REGION Network 11: DB62 DBX3.5 = PIT358 LO / DB62 DBX3.6 = PIT358 HI Fresh Water Inlet Pressure
   // GCU_WARNING_WORD_02_BIT_13
   RUNG wire#powerrail
      "PIT358_ALM_ANALOG_DB78"(Enable := wire#w1, Value := "12_AI_Data".PIT_358_SCALED, "Raw Value" := "Fresh Water Inlet Pressure", "Enable Delay Time" :=, "High Value Release" :=, "SHORT CIRCUIT VALUE" := 32000.0, "BROKEN WIRE VALUE" := -32000.0, "VERY LOW LEVEL VALUE (LL)" := "19_AUTO_CMNDS_Data".PIT358_CMND_LowLow, "LOW LEVEL VALUE (L)" := "19_AUTO_CMNDS_Data".PIT358_CMND_Low, "HIGH LEVEL VALUE (H)" := "19_AUTO_CMNDS_Data".PIT358_CMND_High, "VERY HIGH LEVEL VALUE (HH)" := "19_AUTO_CMNDS_Data".PIT358_CMND_HighHigh, OFFSET :=, "ALARM DELAY" := "86_Times"."PIT358 Delay", "Peak Value Reset" :=, "ALARM HH" =>, "ALARM H" =>, "ALARM L" =>, "ALARM LL" =>, "ALARM READING" => %DB62.DBX1.0, "Peak Value" =>, Alarm =>, Alarm_INT =>)
      wire#w2
      Contact( "10_DI_DATA".P_304_ENBLD )
      wire#w3
      Contact( "PIT358_ALM_ANALOG_DB78"."ALARM L" )
      Coil( %DB62.DBX3.5 )
   END_RUNG
   RUNG wire#powerrail
      { S7_Templates := "SrcType := Int" } GE_Contact(in1 := "100_GCU_AUTO_SEQ_DB".CRNT_STEP, in2 := 140)
      { S7_Templates := "SrcType := Int" } LE_Contact(in1 := "100_GCU_AUTO_SEQ_DB".CRNT_STEP, in2 := 150)
   END_RUNG wire#w1
   RUNG wire#w2
      Contact( "AlwaysTRUE" )
   END_RUNG wire#w3
   RUNG wire#w3
      Contact( "PIT358_ALM_ANALOG_DB78"."ALARM H" )
      Coil( %DB62.DBX3.6 )
   END_RUNG
   // the same network as SCL:
   "PIT358_ALM_ANALOG_DB78"(Value := "12_AI_Data".PIT_358_SCALED,   // "502_ALM_ANALOG"
                           "Raw Value" := "Fresh Water Inlet Pressure",
                           Enable := ("100_GCU_AUTO_SEQ_DB".CRNT_STEP >= 140) AND ("100_GCU_AUTO_SEQ_DB".CRNT_STEP <= 150),
                           "SHORT CIRCUIT VALUE" := 32000.0,
                           "BROKEN WIRE VALUE" := -32000.0,
                           "VERY LOW LEVEL VALUE (LL)" := "19_AUTO_CMNDS_Data".PIT358_CMND_LowLow,
                           "LOW LEVEL VALUE (L)" := "19_AUTO_CMNDS_Data".PIT358_CMND_Low,
                           "HIGH LEVEL VALUE (H)" := "19_AUTO_CMNDS_Data".PIT358_CMND_High,
                           "VERY HIGH LEVEL VALUE (HH)" := "19_AUTO_CMNDS_Data".PIT358_CMND_HighHigh,
                           "ALARM DELAY" := "86_Times"."PIT358 Delay",
                           "ALARM READING" => %DB62.DBX1.0,
                           ENO => #_w1);
   #_w2 := #_w1 AND ("10_DI_DATA".P_304_ENBLD OR "AlwaysTRUE");
   %DB62.DBX3.5 := #_w2 AND "PIT358_ALM_ANALOG_DB78"."ALARM L";
   %DB62.DBX3.6 := #_w2 AND "PIT358_ALM_ANALOG_DB78"."ALARM H";
END_REGION

REGION Network 12: DB62 DBX3.7 = FS350 Fresh Water Cooling Flow Switch
   // GCU_WARNING_WORD_02_BIT_15
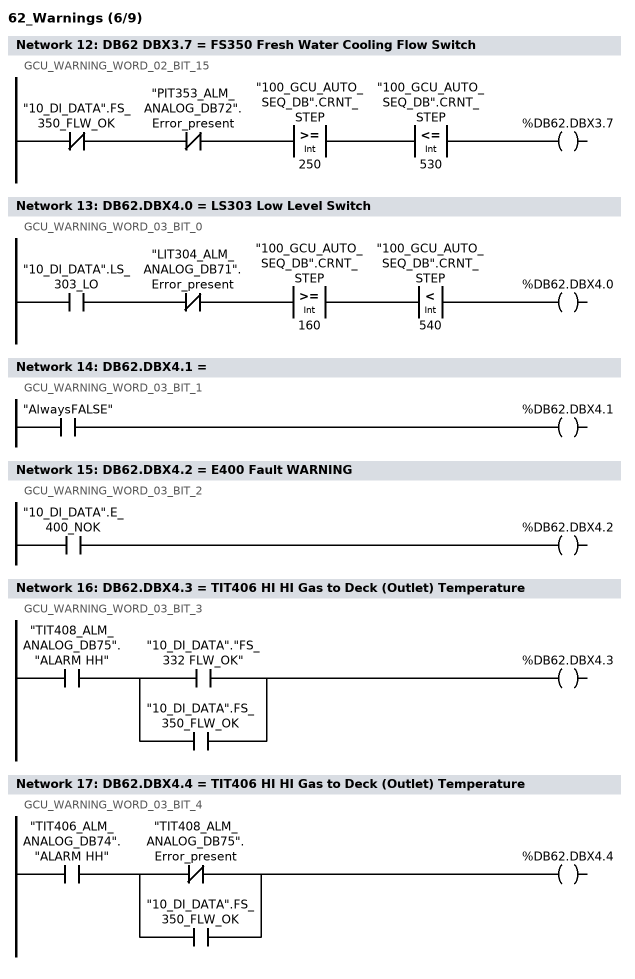
   RUNG wire#powerrail
      I_Contact( "10_DI_DATA".FS_350_FLW_OK )
      I_Contact( "PIT353_ALM_ANALOG_DB72".Error_present )
      { S7_Templates := "SrcType := Int" } GE_Contact(in1 := "100_GCU_AUTO_SEQ_DB".CRNT_STEP, in2 := 250)
      { S7_Templates := "SrcType := Int" } LE_Contact(in1 := "100_GCU_AUTO_SEQ_DB".CRNT_STEP, in2 := 530)
      Coil( %DB62.DBX3.7 )
   END_RUNG
   // the same network as SCL:
   %DB62.DBX3.7 := NOT "10_DI_DATA".FS_350_FLW_OK AND NOT "PIT353_ALM_ANALOG_DB72".Error_present AND ("100_GCU_AUTO_SEQ_DB".CRNT_STEP >= 250) AND ("100_GCU_AUTO_SEQ_DB".CRNT_STEP <= 530);
END_REGION

REGION Network 13: DB62.DBX4.0 = LS303 Low Level Switch
   // GCU_WARNING_WORD_03_BIT_0
   RUNG wire#powerrail
      Contact( "10_DI_DATA".LS_303_LO )
      I_Contact( "LIT304_ALM_ANALOG_DB71".Error_present )
      { S7_Templates := "SrcType := Int" } GE_Contact(in1 := "100_GCU_AUTO_SEQ_DB".CRNT_STEP, in2 := 160)
      { S7_Templates := "SrcType := Int" } LT_Contact(in1 := "100_GCU_AUTO_SEQ_DB".CRNT_STEP, in2 := 540)
      Coil( %DB62.DBX4.0 )
   END_RUNG
   // the same network as SCL:
   %DB62.DBX4.0 := "10_DI_DATA".LS_303_LO AND NOT "LIT304_ALM_ANALOG_DB71".Error_present AND ("100_GCU_AUTO_SEQ_DB".CRNT_STEP >= 160) AND ("100_GCU_AUTO_SEQ_DB".CRNT_STEP < 540);
END_REGION

REGION Network 14: DB62.DBX4.1 =
   // GCU_WARNING_WORD_03_BIT_1
   RUNG wire#powerrail
      Contact( "AlwaysFALSE" )
      Coil( %DB62.DBX4.1 )
   END_RUNG
   // the same network as SCL:
   %DB62.DBX4.1 := "AlwaysFALSE";
END_REGION

REGION Network 15: DB62.DBX4.2 = E400 Fault WARNING
   // GCU_WARNING_WORD_03_BIT_2
   RUNG wire#powerrail
      Contact( "10_DI_DATA".E_400_NOK )
      Coil( %DB62.DBX4.2 )
   END_RUNG
   // the same network as SCL:
   %DB62.DBX4.2 := "10_DI_DATA".E_400_NOK;
END_REGION

REGION Network 16: DB62.DBX4.3 = TIT406 HI HI Gas to Deck (Outlet) Temperature
   // GCU_WARNING_WORD_03_BIT_3
   RUNG wire#powerrail
      Contact( "TIT408_ALM_ANALOG_DB75"."ALARM HH" )
      wire#w1
      Contact( "10_DI_DATA"."FS_332 FLW_OK" )
      wire#w2
      Coil( %DB62.DBX4.3 )
   END_RUNG
   RUNG wire#w1
      Contact( "10_DI_DATA".FS_350_FLW_OK )
   END_RUNG wire#w2
   // the same network as SCL:
   %DB62.DBX4.3 := "TIT408_ALM_ANALOG_DB75"."ALARM HH" AND ("10_DI_DATA"."FS_332 FLW_OK" OR "10_DI_DATA".FS_350_FLW_OK);
END_REGION

REGION Network 17: DB62.DBX4.4 = TIT406 HI HI Gas to Deck (Outlet) Temperature
   // GCU_WARNING_WORD_03_BIT_4
   RUNG wire#powerrail
      Contact( "TIT406_ALM_ANALOG_DB74"."ALARM HH" )
      wire#w1
      I_Contact( "TIT408_ALM_ANALOG_DB75".Error_present )
      wire#w2
      Coil( %DB62.DBX4.4 )
   END_RUNG
   RUNG wire#w1
      Contact( "10_DI_DATA".FS_350_FLW_OK )
   END_RUNG wire#w2
   // the same network as SCL:
   %DB62.DBX4.4 := "TIT406_ALM_ANALOG_DB74"."ALARM HH" AND (NOT "TIT408_ALM_ANALOG_DB75".Error_present OR "10_DI_DATA".FS_350_FLW_OK);
END_REGION

REGION Network 19: New Warning
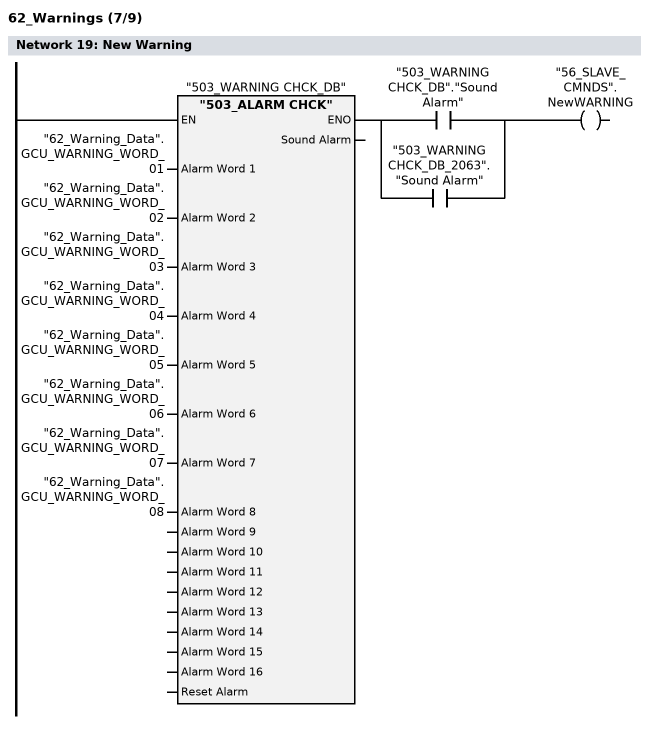
   RUNG wire#powerrail
      "503_WARNING CHCK_DB"("Alarm Word 1" := "62_Warning_Data".GCU_WARNING_WORD_01, "Alarm Word 2" := "62_Warning_Data".GCU_WARNING_WORD_02, "Alarm Word 3" := "62_Warning_Data".GCU_WARNING_WORD_03, "Alarm Word 4" := "62_Warning_Data".GCU_WARNING_WORD_04, "Alarm Word 5" := "62_Warning_Data".GCU_WARNING_WORD_05, "Alarm Word 6" := "62_Warning_Data".GCU_WARNING_WORD_06, "Alarm Word 7" := "62_Warning_Data".GCU_WARNING_WORD_07, "Alarm Word 8" := "62_Warning_Data".GCU_WARNING_WORD_08, "Alarm Word 9" :=, "Alarm Word 10" :=, "Alarm Word 11" :=, "Alarm Word 12" :=, "Alarm Word 13" :=, "Alarm Word 14" :=, "Alarm Word 15" :=, "Alarm Word 16" :=, "Reset Alarm" :=, "Sound Alarm" =>)
      wire#w1
      Contact( "503_WARNING CHCK_DB"."Sound Alarm" )
      wire#w2
      Coil( "56_SLAVE_CMNDS".NewWARNING )
   END_RUNG
   RUNG wire#w1
      Contact( "503_WARNING CHCK_DB_2063"."Sound Alarm" )
   END_RUNG wire#w2
   // the same network as SCL:
   "503_WARNING CHCK_DB"("Alarm Word 1" := "62_Warning_Data".GCU_WARNING_WORD_01,   // "503_ALARM CHCK"
                         "Alarm Word 2" := "62_Warning_Data".GCU_WARNING_WORD_02,
                         "Alarm Word 3" := "62_Warning_Data".GCU_WARNING_WORD_03,
                         "Alarm Word 4" := "62_Warning_Data".GCU_WARNING_WORD_04,
                         "Alarm Word 5" := "62_Warning_Data".GCU_WARNING_WORD_05,
                         "Alarm Word 6" := "62_Warning_Data".GCU_WARNING_WORD_06,
                         "Alarm Word 7" := "62_Warning_Data".GCU_WARNING_WORD_07,
                         "Alarm Word 8" := "62_Warning_Data".GCU_WARNING_WORD_08,
                         ENO => #_w1);
   "56_SLAVE_CMNDS".NewWARNING := #_w1 AND ("503_WARNING CHCK_DB"."Sound Alarm" OR "503_WARNING CHCK_DB_2063"."Sound Alarm");
END_REGION

REGION Network 20: Warning Present
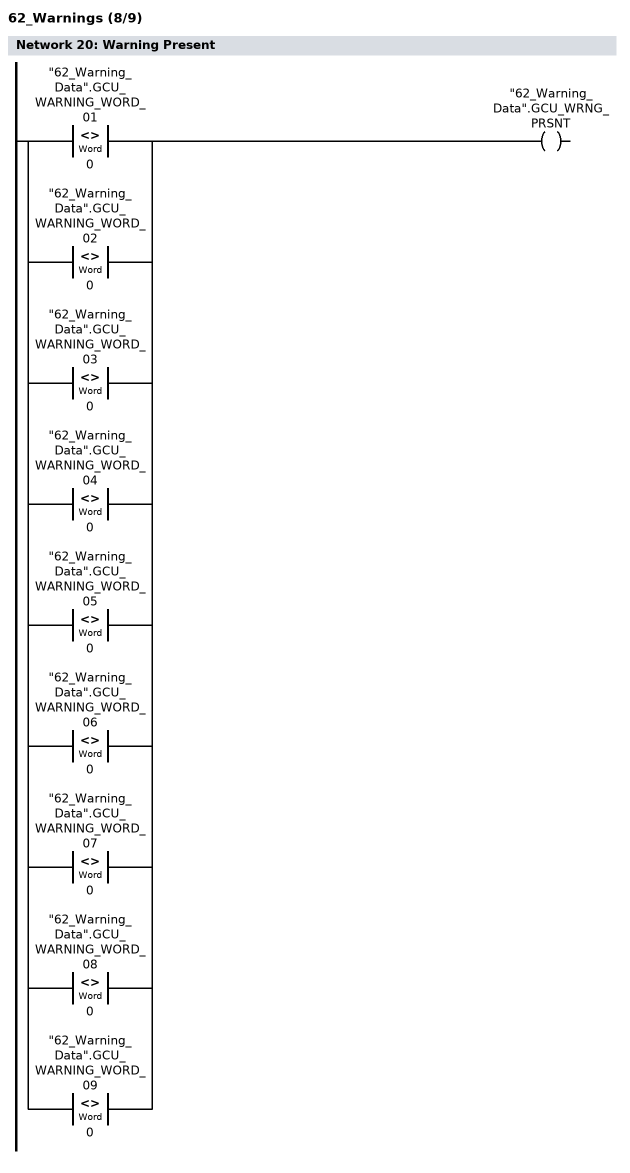
   RUNG wire#powerrail
      { S7_Templates := "SrcType := Word" } NE_Contact(in1 := "62_Warning_Data".GCU_WARNING_WORD_01, in2 := 0)
      wire#w1
      Coil( "62_Warning_Data".GCU_WRNG_PRSNT )
   END_RUNG
   RUNG wire#powerrail
      { S7_Templates := "SrcType := Word" } NE_Contact(in1 := "62_Warning_Data".GCU_WARNING_WORD_02, in2 := 0)
   END_RUNG wire#w1
   RUNG wire#powerrail
      { S7_Templates := "SrcType := Word" } NE_Contact(in1 := "62_Warning_Data".GCU_WARNING_WORD_03, in2 := 0)
   END_RUNG wire#w1
   RUNG wire#powerrail
      { S7_Templates := "SrcType := Word" } NE_Contact(in1 := "62_Warning_Data".GCU_WARNING_WORD_04, in2 := 0)
   END_RUNG wire#w1
   RUNG wire#powerrail
      { S7_Templates := "SrcType := Word" } NE_Contact(in1 := "62_Warning_Data".GCU_WARNING_WORD_05, in2 := 0)
   END_RUNG wire#w1
   RUNG wire#powerrail
      { S7_Templates := "SrcType := Word" } NE_Contact(in1 := "62_Warning_Data".GCU_WARNING_WORD_06, in2 := 0)
   END_RUNG wire#w1
   RUNG wire#powerrail
      { S7_Templates := "SrcType := Word" } NE_Contact(in1 := "62_Warning_Data".GCU_WARNING_WORD_07, in2 := 0)
   END_RUNG wire#w1
   RUNG wire#powerrail
      { S7_Templates := "SrcType := Word" } NE_Contact(in1 := "62_Warning_Data".GCU_WARNING_WORD_08, in2 := 0)
   END_RUNG wire#w1
   RUNG wire#powerrail
      { S7_Templates := "SrcType := Word" } NE_Contact(in1 := "62_Warning_Data".GCU_WARNING_WORD_09, in2 := 0)
   END_RUNG wire#w1
   // the same network as SCL:
   "62_Warning_Data".GCU_WRNG_PRSNT := ("62_Warning_Data".GCU_WARNING_WORD_01 <> 0) OR ("62_Warning_Data".GCU_WARNING_WORD_02 <> 0) OR ("62_Warning_Data".GCU_WARNING_WORD_03 <> 0) OR ("62_Warning_Data".GCU_WARNING_WORD_04 <> 0) OR ("62_Warning_Data".GCU_WARNING_WORD_05 <> 0) OR ("62_Warning_Data".GCU_WARNING_WORD_06 <> 0) OR ("62_Warning_Data".GCU_WARNING_WORD_07 <> 0) OR ("62_Warning_Data".GCU_WARNING_WORD_08 <> 0) OR ("62_Warning_Data".GCU_WARNING_WORD_09 <> 0);
END_REGION

REGION Network 21: Master Warning
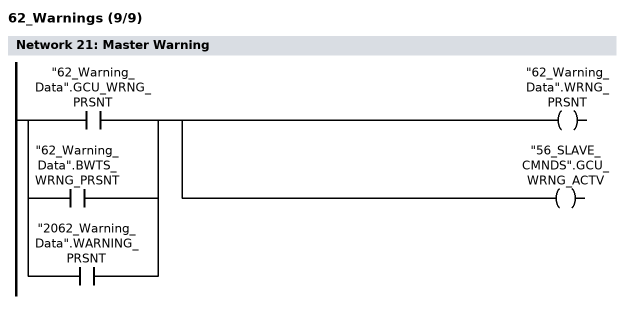
   RUNG wire#powerrail
      Contact( "62_Warning_Data".GCU_WRNG_PRSNT )
      wire#w1
      Coil( "62_Warning_Data".WRNG_PRSNT )
   END_RUNG
   RUNG wire#powerrail
      Contact( "62_Warning_Data".BWTS_WRNG_PRSNT )
   END_RUNG wire#w1
   RUNG wire#powerrail
      Contact( "2062_Warning_Data".WARNING_PRSNT )
   END_RUNG wire#w1
   RUNG wire#w1
      Coil( "56_SLAVE_CMNDS".GCU_WRNG_ACTV )
   END_RUNG
   // the same network as SCL:
   "62_Warning_Data".WRNG_PRSNT := "62_Warning_Data".GCU_WRNG_PRSNT OR "62_Warning_Data".BWTS_WRNG_PRSNT OR "2062_Warning_Data".WARNING_PRSNT;
   "56_SLAVE_CMNDS".GCU_WRNG_ACTV := "62_Warning_Data".WRNG_PRSNT;
END_REGION
END_FUNCTION

FUNCTION "68_Sys_Status" : Void   // FC68, LAD
TITLE = System Status
{ S7_Optimized_Access := 'TRUE' }
AUTHOR : JRS
VERSION : 0.1
// For the determination of specific system status information as required by the code
   VAR_TEMP   // added for the SCL form of the ladder/FBD networks
      _w1 : Bool;
   END_VAR
BEGIN

REGION Network 1: Valves At Initial
   // All valves in initial state
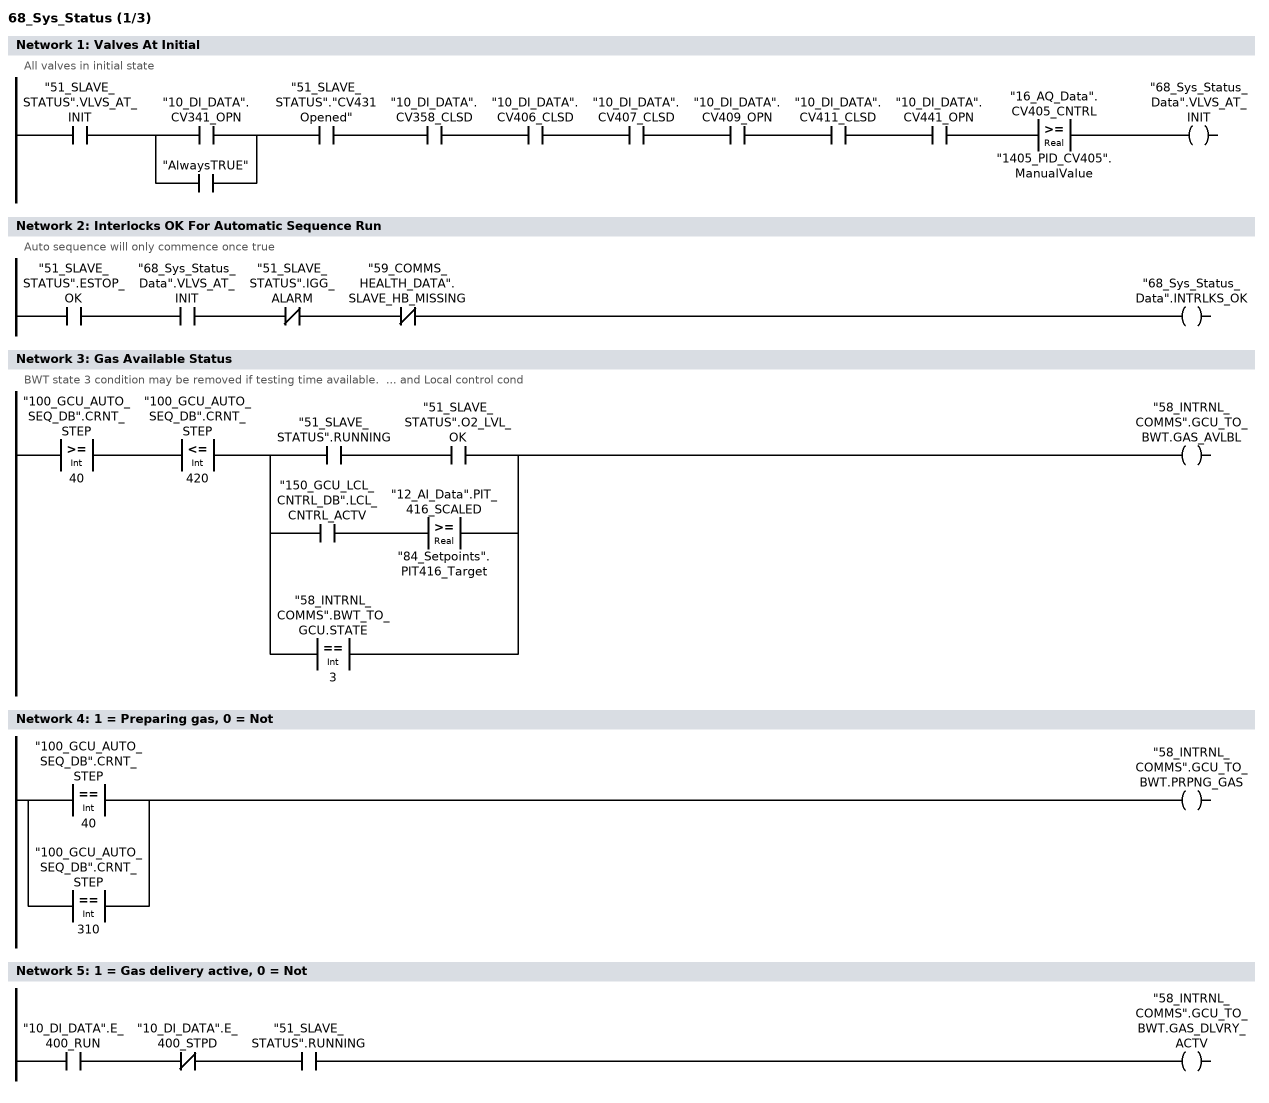
   RUNG wire#powerrail
      Contact( "51_SLAVE_STATUS".VLVS_AT_INIT )
      wire#w1
      Contact( "10_DI_DATA".CV341_OPN )
      wire#w2
      Contact( "51_SLAVE_STATUS"."CV431 Opened" )
      Contact( "10_DI_DATA".CV358_CLSD )
      Contact( "10_DI_DATA".CV406_CLSD )
      Contact( "10_DI_DATA".CV407_CLSD )
      Contact( "10_DI_DATA".CV409_OPN )
      Contact( "10_DI_DATA".CV411_CLSD )
      Contact( "10_DI_DATA".CV441_OPN )
      { S7_Templates := "SrcType := Real" } GE_Contact(in1 := "16_AQ_Data".CV405_CNTRL, in2 := "1405_PID_CV405".ManualValue)
      Coil( "68_Sys_Status_Data".VLVS_AT_INIT )
   END_RUNG
   RUNG wire#w1
      Contact( "AlwaysTRUE" )
   END_RUNG wire#w2
   // the same network as SCL:
   "68_Sys_Status_Data".VLVS_AT_INIT := "51_SLAVE_STATUS".VLVS_AT_INIT AND ("10_DI_DATA".CV341_OPN OR "AlwaysTRUE") AND "51_SLAVE_STATUS"."CV431 Opened" AND "10_DI_DATA".CV358_CLSD AND "10_DI_DATA".CV406_CLSD AND "10_DI_DATA".CV407_CLSD AND "10_DI_DATA".CV409_OPN AND "10_DI_DATA".CV411_CLSD AND "10_DI_DATA".CV441_OPN AND ("16_AQ_Data".CV405_CNTRL >= "1405_PID_CV405".ManualValue);
END_REGION

REGION Network 2: Interlocks OK For Automatic Sequence Run
   // Auto sequence will only commence once true
   RUNG wire#powerrail
      Contact( "51_SLAVE_STATUS".ESTOP_OK )
      Contact( "68_Sys_Status_Data".VLVS_AT_INIT )
      I_Contact( "51_SLAVE_STATUS".IGG_ALARM )
      I_Contact( "59_COMMS_HEALTH_DATA".SLAVE_HB_MISSING )
      Coil( "68_Sys_Status_Data".INTRLKS_OK )
   END_RUNG
   // the same network as SCL:
   "68_Sys_Status_Data".INTRLKS_OK := "51_SLAVE_STATUS".ESTOP_OK AND "68_Sys_Status_Data".VLVS_AT_INIT AND NOT "51_SLAVE_STATUS".IGG_ALARM AND NOT "59_COMMS_HEALTH_DATA".SLAVE_HB_MISSING;
END_REGION

REGION Network 3: Gas Available Status
   // BWT state 3 condition may be removed if testing time available.  ... and Local control cond
   RUNG wire#powerrail
      { S7_Templates := "SrcType := Int" } GE_Contact(in1 := "100_GCU_AUTO_SEQ_DB".CRNT_STEP, in2 := 40)
      { S7_Templates := "SrcType := Int" } LE_Contact(in1 := "100_GCU_AUTO_SEQ_DB".CRNT_STEP, in2 := 420)
      wire#w1
      Contact( "51_SLAVE_STATUS".RUNNING )
      Contact( "51_SLAVE_STATUS".O2_LVL_OK )
      wire#w2
      Coil( "58_INTRNL_COMMS".GCU_TO_BWT.GAS_AVLBL )
   END_RUNG
   RUNG wire#w1
      Contact( "150_GCU_LCL_CNTRL_DB".LCL_CNTRL_ACTV )
      { S7_Templates := "SrcType := Real" } GE_Contact(in1 := "12_AI_Data".PIT_416_SCALED, in2 := "84_Setpoints".PIT416_Target)
   END_RUNG wire#w2
   RUNG wire#w1
      { S7_Templates := "SrcType := Int" } EQ_Contact(in1 := "58_INTRNL_COMMS".BWT_TO_GCU.STATE, in2 := 3)
   END_RUNG wire#w2
   // the same network as SCL:
   "58_INTRNL_COMMS".GCU_TO_BWT.GAS_AVLBL := ("100_GCU_AUTO_SEQ_DB".CRNT_STEP >= 40) AND ("100_GCU_AUTO_SEQ_DB".CRNT_STEP <= 420) AND (("51_SLAVE_STATUS".RUNNING AND "51_SLAVE_STATUS".O2_LVL_OK) OR ("150_GCU_LCL_CNTRL_DB".LCL_CNTRL_ACTV AND ("12_AI_Data".PIT_416_SCALED >= "84_Setpoints".PIT416_Target)) OR ("58_INTRNL_COMMS".BWT_TO_GCU.STATE = 3));
END_REGION

REGION Network 4: 1 = Preparing gas, 0 = Not
   RUNG wire#powerrail
      { S7_Templates := "SrcType := Int" } EQ_Contact(in1 := "100_GCU_AUTO_SEQ_DB".CRNT_STEP, in2 := 40)
      wire#w1
      Coil( "58_INTRNL_COMMS".GCU_TO_BWT.PRPNG_GAS )
   END_RUNG
   RUNG wire#powerrail
      { S7_Templates := "SrcType := Int" } EQ_Contact(in1 := "100_GCU_AUTO_SEQ_DB".CRNT_STEP, in2 := 310)
   END_RUNG wire#w1
   // the same network as SCL:
   "58_INTRNL_COMMS".GCU_TO_BWT.PRPNG_GAS := ("100_GCU_AUTO_SEQ_DB".CRNT_STEP = 40) OR ("100_GCU_AUTO_SEQ_DB".CRNT_STEP = 310);
END_REGION

REGION Network 5: 1 = Gas delivery active, 0 = Not
   RUNG wire#powerrail
      Contact( "10_DI_DATA".E_400_RUN )
      I_Contact( "10_DI_DATA".E_400_STPD )
      Contact( "51_SLAVE_STATUS".RUNNING )
      Coil( "58_INTRNL_COMMS".GCU_TO_BWT.GAS_DLVRY_ACTV )
   END_RUNG
   // the same network as SCL:
   "58_INTRNL_COMMS".GCU_TO_BWT.GAS_DLVRY_ACTV := "10_DI_DATA".E_400_RUN AND NOT "10_DI_DATA".E_400_STPD AND "51_SLAVE_STATUS".RUNNING;
END_REGION

REGION Network 6: PGC Hours Run
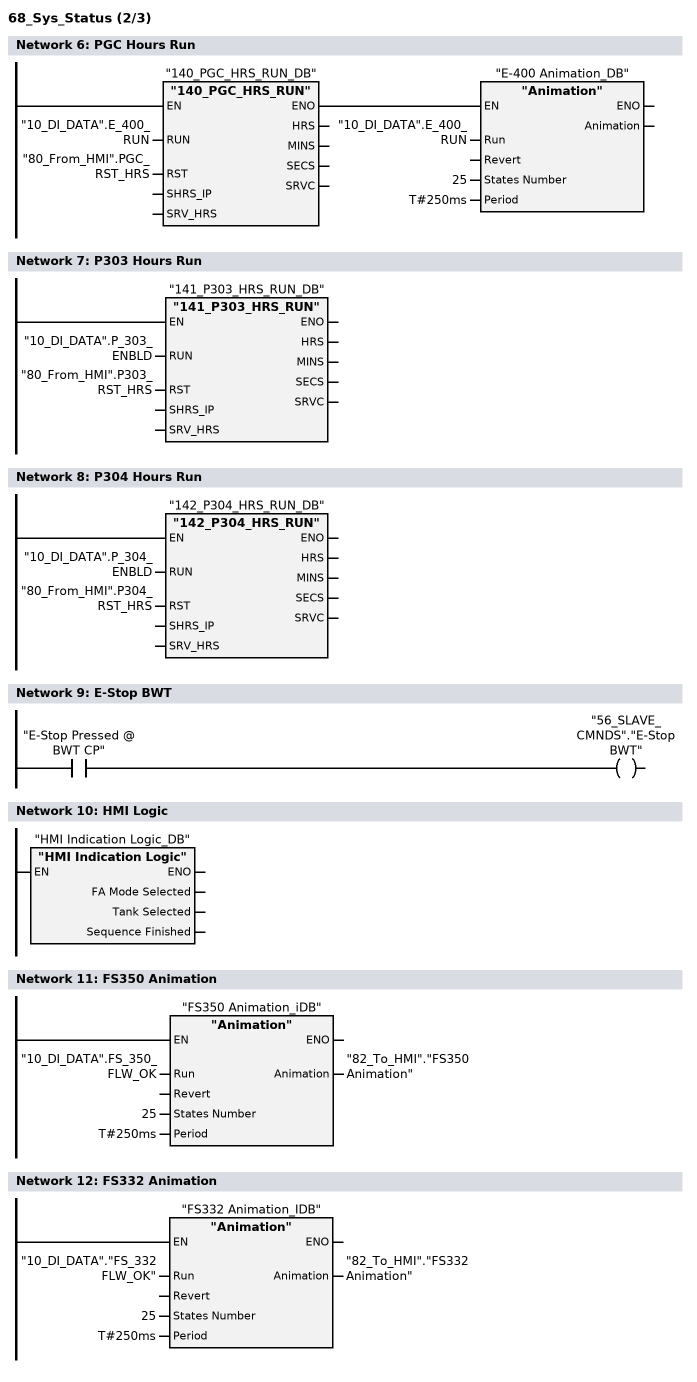
   RUNG wire#powerrail
      "140_PGC_HRS_RUN_DB"(RUN := "10_DI_DATA".E_400_RUN, RST := "80_From_HMI".PGC_RST_HRS, SHRS_IP :=, SRV_HRS :=, HRS =>, MINS =>, SECS =>, SRVC =>)
      "E-400 Animation_DB"(Run := "10_DI_DATA".E_400_RUN, Revert :=, "States Number" := 25, Period := T#250ms, Animation =>)
   END_RUNG
   // the same network as SCL:
   "140_PGC_HRS_RUN_DB"(RUN := "10_DI_DATA".E_400_RUN, RST := "80_From_HMI".PGC_RST_HRS, ENO => #_w1);   // "140_PGC_HRS_RUN"
   IF #_w1 THEN
       "E-400 Animation_DB"(Run := "10_DI_DATA".E_400_RUN, "States Number" := 25, Period := T#250ms);   // "Animation"
   END_IF;
END_REGION

REGION Network 7: P303 Hours Run
   RUNG wire#powerrail
      "141_P303_HRS_RUN_DB"(RUN := "10_DI_DATA".P_303_ENBLD, RST := "80_From_HMI".P303_RST_HRS, SHRS_IP :=, SRV_HRS :=, HRS =>, MINS =>, SECS =>, SRVC =>)
   END_RUNG
   // the same network as SCL:
   "141_P303_HRS_RUN_DB"(RUN := "10_DI_DATA".P_303_ENBLD, RST := "80_From_HMI".P303_RST_HRS);   // "141_P303_HRS_RUN"
END_REGION

REGION Network 8: P304 Hours Run
   RUNG wire#powerrail
      "142_P304_HRS_RUN_DB"(RUN := "10_DI_DATA".P_304_ENBLD, RST := "80_From_HMI".P304_RST_HRS, SHRS_IP :=, SRV_HRS :=, HRS =>, MINS =>, SECS =>, SRVC =>)
   END_RUNG
   // the same network as SCL:
   "142_P304_HRS_RUN_DB"(RUN := "10_DI_DATA".P_304_ENBLD, RST := "80_From_HMI".P304_RST_HRS);   // "142_P304_HRS_RUN"
END_REGION

REGION Network 9: E-Stop BWT
   RUNG wire#powerrail
      Contact( "E-Stop Pressed @ BWT CP" )
      Coil( "56_SLAVE_CMNDS"."E-Stop BWT" )
   END_RUNG
   // the same network as SCL:
   "56_SLAVE_CMNDS"."E-Stop BWT" := "E-Stop Pressed @ BWT CP";
END_REGION

REGION Network 10: HMI Logic
   RUNG wire#powerrail
      "HMI Indication Logic_DB"("FA Mode Selected" =>, "Tank Selected" =>, "Sequence Finished" =>)
   END_RUNG
   // the same network as SCL:
   "HMI Indication Logic_DB"();   // "HMI Indication Logic"
END_REGION

REGION Network 11: FS350 Animation
   RUNG wire#powerrail
      "FS350 Animation_iDB"(Run := "10_DI_DATA".FS_350_FLW_OK, Revert :=, "States Number" := 25, Period := T#250ms, Animation => "82_To_HMI"."FS350 Animation")
   END_RUNG
   // the same network as SCL:
   "FS350 Animation_iDB"(Run := "10_DI_DATA".FS_350_FLW_OK,   // "Animation"
                         "States Number" := 25,
                         Period := T#250ms,
                         Animation => "82_To_HMI"."FS350 Animation");
END_REGION

REGION Network 12: FS332 Animation
   RUNG wire#powerrail
      "FS332 Animation_IDB"(Run := "10_DI_DATA"."FS_332 FLW_OK", Revert :=, "States Number" := 25, Period := T#250ms, Animation => "82_To_HMI"."FS332 Animation")
   END_RUNG
   // the same network as SCL:
   "FS332 Animation_IDB"(Run := "10_DI_DATA"."FS_332 FLW_OK",   // "Animation"
                         "States Number" := 25,
                         Period := T#250ms,
                         Animation => "82_To_HMI"."FS332 Animation");
END_REGION

REGION Network 13: FS332 Animation
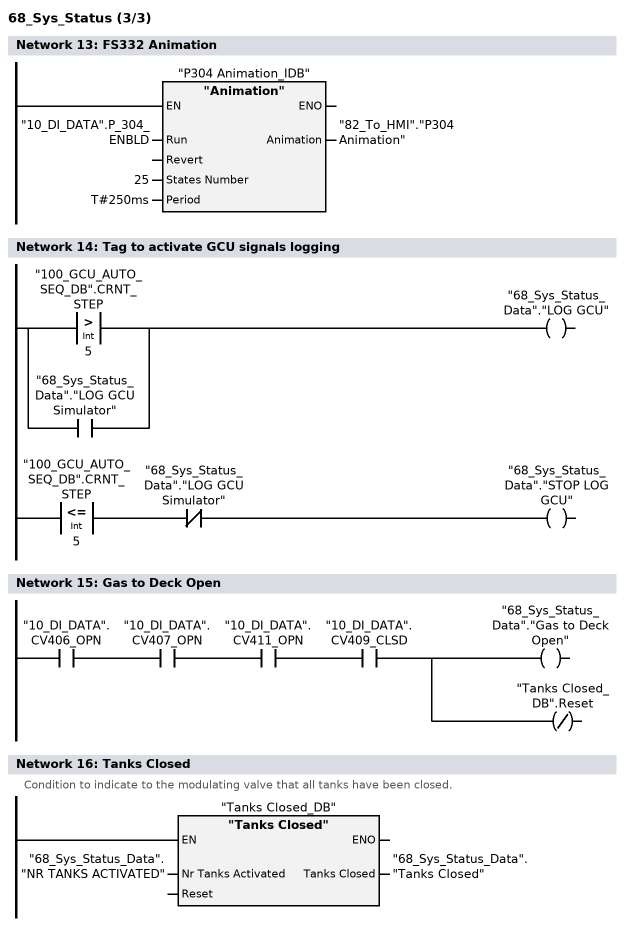
   RUNG wire#powerrail
      "P304 Animation_IDB"(Run := "10_DI_DATA".P_304_ENBLD, Revert :=, "States Number" := 25, Period := T#250ms, Animation => "82_To_HMI"."P304 Animation")
   END_RUNG
   // the same network as SCL:
   "P304 Animation_IDB"(Run := "10_DI_DATA".P_304_ENBLD,   // "Animation"
                        "States Number" := 25,
                        Period := T#250ms,
                        Animation => "82_To_HMI"."P304 Animation");
END_REGION

REGION Network 14: Tag to activate GCU signals logging
   RUNG wire#powerrail
      { S7_Templates := "SrcType := Int" } GT_Contact(in1 := "100_GCU_AUTO_SEQ_DB".CRNT_STEP, in2 := 5)
      wire#w1
      Coil( "68_Sys_Status_Data"."LOG GCU" )
   END_RUNG
   RUNG wire#powerrail
      Contact( "68_Sys_Status_Data"."LOG GCU Simulator" )
   END_RUNG wire#w1
   RUNG wire#powerrail
      { S7_Templates := "SrcType := Int" } LE_Contact(in1 := "100_GCU_AUTO_SEQ_DB".CRNT_STEP, in2 := 5)
      I_Contact( "68_Sys_Status_Data"."LOG GCU Simulator" )
      Coil( "68_Sys_Status_Data"."STOP LOG GCU" )
   END_RUNG
   // the same network as SCL:
   "68_Sys_Status_Data"."LOG GCU" := ("100_GCU_AUTO_SEQ_DB".CRNT_STEP > 5) OR "68_Sys_Status_Data"."LOG GCU Simulator";
   "68_Sys_Status_Data"."STOP LOG GCU" := ("100_GCU_AUTO_SEQ_DB".CRNT_STEP <= 5) AND NOT "68_Sys_Status_Data"."LOG GCU Simulator";
END_REGION

REGION Network 15: Gas to Deck Open
   RUNG wire#powerrail
      Contact( "10_DI_DATA".CV406_OPN )
      Contact( "10_DI_DATA".CV407_OPN )
      Contact( "10_DI_DATA".CV411_OPN )
      Contact( "10_DI_DATA".CV409_CLSD )
      wire#w1
      Coil( "68_Sys_Status_Data"."Gas to Deck Open" )
   END_RUNG
   RUNG wire#w1
      I_Coil( "Tanks Closed_DB".Reset )
   END_RUNG
   // the same network as SCL:
   "68_Sys_Status_Data"."Gas to Deck Open" := "10_DI_DATA".CV406_OPN AND "10_DI_DATA".CV407_OPN AND "10_DI_DATA".CV411_OPN AND "10_DI_DATA".CV409_CLSD;
   "Tanks Closed_DB".Reset := NOT "68_Sys_Status_Data"."Gas to Deck Open";
END_REGION

REGION Network 16: Tanks Closed
   // Condition to indicate to the modulating valve that all tanks have been closed.
   RUNG wire#powerrail
      "Tanks Closed_DB"("Nr Tanks Activated" := "68_Sys_Status_Data"."NR TANKS ACTIVATED", Reset :=, "Tanks Closed" => "68_Sys_Status_Data"."Tanks Closed")
   END_RUNG
   // the same network as SCL:
   "Tanks Closed_DB"("Nr Tanks Activated" := "68_Sys_Status_Data"."NR TANKS ACTIVATED",   // "Tanks Closed"
                     "Tanks Closed" => "68_Sys_Status_Data"."Tanks Closed");
END_REGION
END_FUNCTION

// folder: 70 - 79 Modes of Operation

FUNCTION "70_Mode_Control" : Void   // FC70, LAD
TITLE = Mode Control
{ S7_Optimized_Access := 'TRUE' }
AUTHOR : JRS
VERSION : 0.1
// To determine the current mode of operation 1=Auto(default), 2=Manual, 3=FatAuto, 4=FatManual
   VAR_TEMP   // added for the SCL form of the ladder/FBD networks
      _w1 : Bool;
   END_VAR
BEGIN

REGION Network 1: Default = Automatic
   // Set default to Automatic (on first scan)
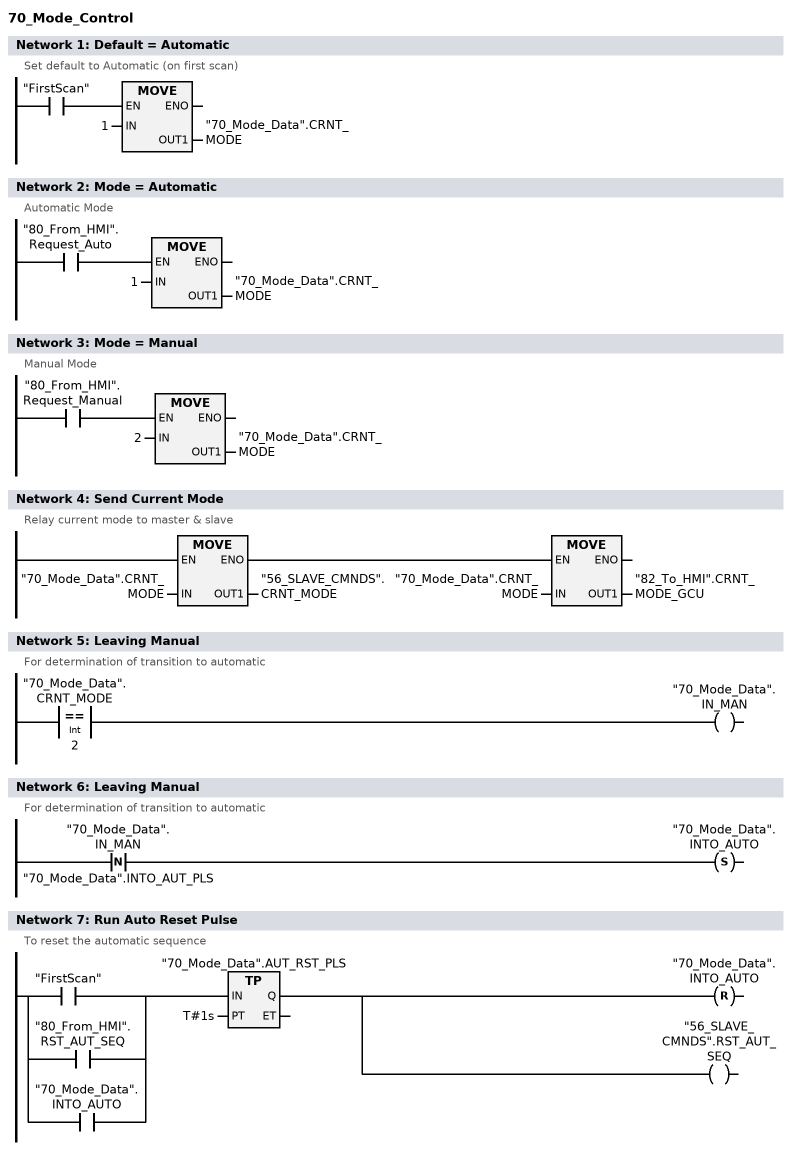
   RUNG wire#powerrail
      Contact( "FirstScan" )
      Move(in := 1, out1 => "70_Mode_Data".CRNT_MODE)
   END_RUNG
   // the same network as SCL:
   IF "FirstScan" THEN "70_Mode_Data".CRNT_MODE := 1; END_IF;
END_REGION

REGION Network 2: Mode = Automatic
   // Automatic Mode
   RUNG wire#powerrail
      Contact( "80_From_HMI".Request_Auto )
      Move(in := 1, out1 => "70_Mode_Data".CRNT_MODE)
   END_RUNG
   // the same network as SCL:
   IF "80_From_HMI".Request_Auto THEN "70_Mode_Data".CRNT_MODE := 1; END_IF;
END_REGION

REGION Network 3: Mode = Manual
   // Manual Mode
   RUNG wire#powerrail
      Contact( "80_From_HMI".Request_Manual )
      Move(in := 2, out1 => "70_Mode_Data".CRNT_MODE)
   END_RUNG
   // the same network as SCL:
   IF "80_From_HMI".Request_Manual THEN "70_Mode_Data".CRNT_MODE := 2; END_IF;
END_REGION

REGION Network 4: Send Current Mode
   // Relay current mode to master & slave
   RUNG wire#powerrail
      Move(in := "70_Mode_Data".CRNT_MODE, out1 => "56_SLAVE_CMNDS".CRNT_MODE)
      Move(in := "70_Mode_Data".CRNT_MODE, out1 => "82_To_HMI".CRNT_MODE_GCU)
   END_RUNG
   // the same network as SCL:
   "56_SLAVE_CMNDS".CRNT_MODE := "70_Mode_Data".CRNT_MODE;
   "82_To_HMI".CRNT_MODE_GCU := "70_Mode_Data".CRNT_MODE;
END_REGION

REGION Network 5: Leaving Manual
   // For determination of transition to automatic
   RUNG wire#powerrail
      { S7_Templates := "SrcType := Int" } EQ_Contact(in1 := "70_Mode_Data".CRNT_MODE, in2 := 2)
      Coil( "70_Mode_Data".IN_MAN )
   END_RUNG
   // the same network as SCL:
   "70_Mode_Data".IN_MAN := "70_Mode_Data".CRNT_MODE = 2;
END_REGION

REGION Network 6: Leaving Manual
   // For determination of transition to automatic
   RUNG wire#powerrail
      N_Contact(operand := "70_Mode_Data".IN_MAN, bit := "70_Mode_Data".INTO_AUT_PLS)
      S_Coil( "70_Mode_Data".INTO_AUTO )
   END_RUNG
   // the same network as SCL:
   #_w1 := NOT "70_Mode_Data".IN_MAN AND "70_Mode_Data".INTO_AUT_PLS;   // falling edge of "70_Mode_Data".IN_MAN
   "70_Mode_Data".INTO_AUT_PLS := "70_Mode_Data".IN_MAN;
   IF #_w1 THEN "70_Mode_Data".INTO_AUTO := TRUE; END_IF;
END_REGION

REGION Network 7: Run Auto Reset Pulse
   // To reset the automatic sequence
   "70_Mode_Data".AUT_RST_PLS.TP(IN := "FirstScan" OR "80_From_HMI".RST_AUT_SEQ OR "70_Mode_Data".INTO_AUTO,
                           PT := T#1s);
   IF "70_Mode_Data".AUT_RST_PLS.Q THEN "70_Mode_Data".INTO_AUTO := FALSE; END_IF;
   "56_SLAVE_CMNDS".RST_AUT_SEQ := "70_Mode_Data".AUT_RST_PLS.Q;
END_REGION
END_FUNCTION

// folder: 80 - 89 HMI Handling

FUNCTION "PGC_COMMISSION_MODE" : Void   // FC1, LAD
{ S7_Optimized_Access := 'TRUE' }
VERSION : 0.1
   VAR_TEMP   // added for the SCL form of the ladder/FBD networks
      _w1 : Bool;
   END_VAR
BEGIN

REGION Network 1: When button pressed write temporary setpoint in